(* Logix 5000 project; controller FV vendor 1 type 14 code 217 rev 31.11; software revision 31.00; part 41 of 63 *)
(* tags used below, declared in another part *)
   CWD : CHECKWORD_FLAGS;
   FV_AV1 : PlantItem;   // AV1
   FV_B100 : INT[255];   // FV FLAGS
   FV_B22 : INT[255];   // YSVFILL_FL YSV filling process flags
   FV_B22_0_2_OutputBit : BOOL;
   fv_data_file_value_to_move : DINT;
   FV_indirect_address : DINT;
   FV_N101 : INT[255];   // FV INT Fermentation control integer workspace
   FV_N104 : INT[255];   // FV_PC_BUF PC>PLC Fermentation Control Command Buff er File
   FV_N12 : INT[255];   // SYS_PARMS System Parameter Fil e
   FV_N141 : INT[255];   // YSV1 DATA
   FV_N142 : INT[255];   // YSV2 DATA
   FV_N143 : INT[255];   // YSV3 DATA
   FV_N144 : INT[255];   // YST1 DATA
   FV_N145 : INT[255];   // YST2 DATA
   FV_N20 : INT[255];   // YSVFILL<PC YSV Filling data fro m PC
   FV_N21 : INT[255];   // YSVFILL>PC YSV Filling process data to PC and contr ol regs
   FV_N24 : INT[255];   // YSVFILL_SV YSV filling process data save file to PC
   FV_YSV2O : PlantItem;   // YSV2O
   FV_YSV3O : PlantItem;   // YSV3O
   indirect_bit_temp : INT;
   YSVFilling_transaction_log_delay : DINT;
(* FV_Common, continued *)

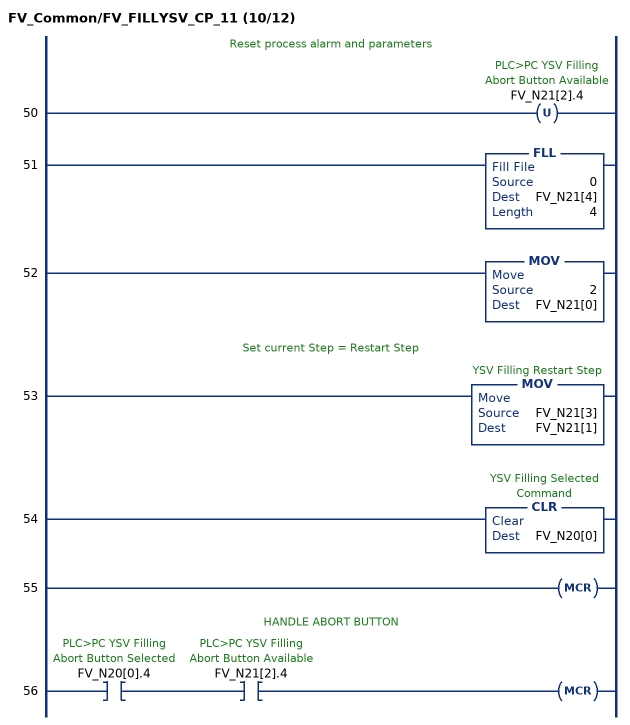
   // Reset process alarm and parameters
   50: OTU(FV_N21[2].4);
   51: FLL(0,FV_N21[4],4);
   52: MOV(2,FV_N21[0]);
   // Set current Step = Restart Step
   53: MOV(FV_N21[3],FV_N21[1]);
   54: CLR(FV_N20[0]);
   55: MCR();
   // HANDLE ABORT BUTTON
   56: XIC(FV_N20[0].4)XIC(FV_N21[2].4)MCR();
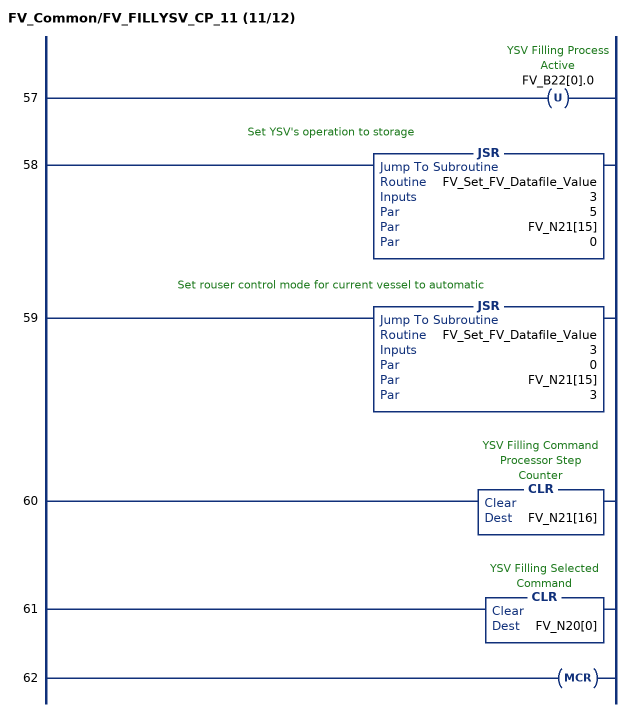
   57: OTU(FV_B22[0].0);
   // Set YSV's operation to storage
   58: JSR(FV_Set_FV_Datafile_Value,3,5,FV_N21[15],0);
   // Set rouser control mode for current vessel to automatic
   59: JSR(FV_Set_FV_Datafile_Value,3,0,FV_N21[15],3);
   60: CLR(FV_N21[16]);
   61: CLR(FV_N20[0]);
   62: MCR();
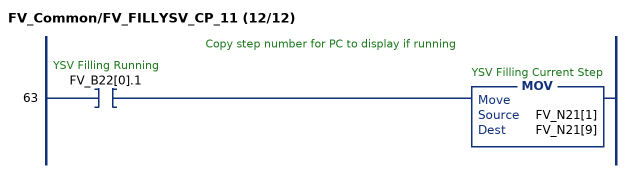
   // Copy step number for PC to display if running
   63: XIC(FV_B22[0].1)MOV(FV_N21[1],FV_N21[9]);
END_ROUTINE

ROUTINE FV_FILLYSV_MC_10   (* ladder *)
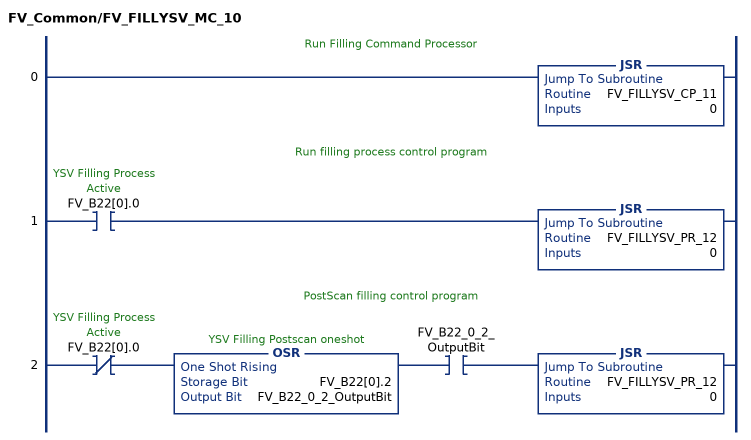
   // Run Filling Command Processor
   0: JSR(FV_FILLYSV_CP_11,0);
   // Run filling process control program
   1: XIC(FV_B22[0].0)JSR(FV_FILLYSV_PR_12,0);
   // PostScan filling control program
   2: XIO(FV_B22[0].0)OSR(FV_B22[0].2,FV_B22_0_2_OutputBit)XIC(FV_B22_0_2_OutputBit)JSR(FV_FILLYSV_PR_12,0);
END_ROUTINE

ROUTINE FV_FILLYSV_PR_12   (* ladder *)
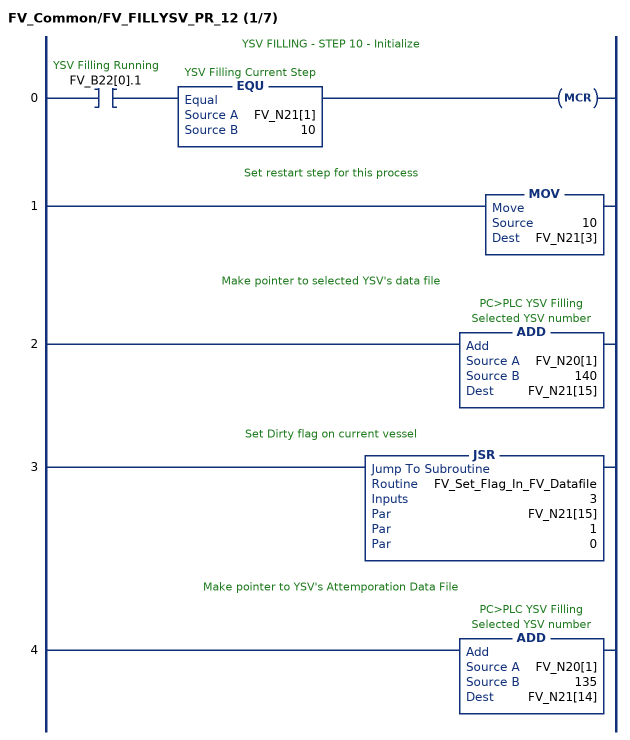
   // YSV FILLING - STEP 10 - Initialize
   0: XIC(FV_B22[0].1)EQU(FV_N21[1],10)MCR();
   // Set restart step for this process
   1: MOV(10,FV_N21[3]);
   // Make pointer to selected YSV's data file
   2: ADD(FV_N20[1],140,FV_N21[15]);
   // Set Dirty flag on current vessel
   3: JSR(FV_Set_Flag_In_FV_Datafile,3,FV_N21[15],1,0);
   // Make pointer to YSV's Attemporation Data File
   4: ADD(FV_N20[1],135,FV_N21[14]);
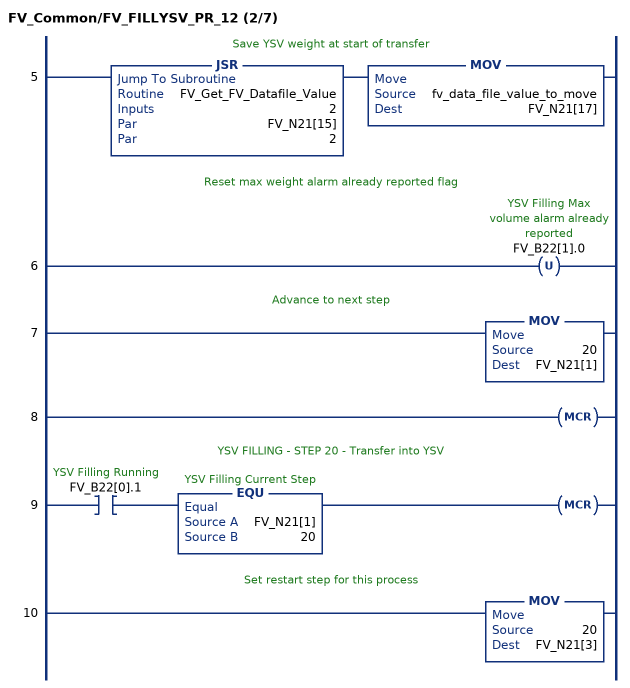
   // Save YSV weight at start of transfer
   5: JSR(FV_Get_FV_Datafile_Value,2,FV_N21[15],2)MOV(fv_data_file_value_to_move,FV_N21[17]);
   // Reset max weight alarm already reported flag
   6: OTU(FV_B22[1].0);
   // Advance to next step
   7: MOV(20,FV_N21[1]);
   8: MCR();
   // YSV FILLING - STEP 20 - Transfer into YSV
   9: XIC(FV_B22[0].1)EQU(FV_N21[1],20)MCR();
   // Set restart step for this process
   10: MOV(20,FV_N21[3]);
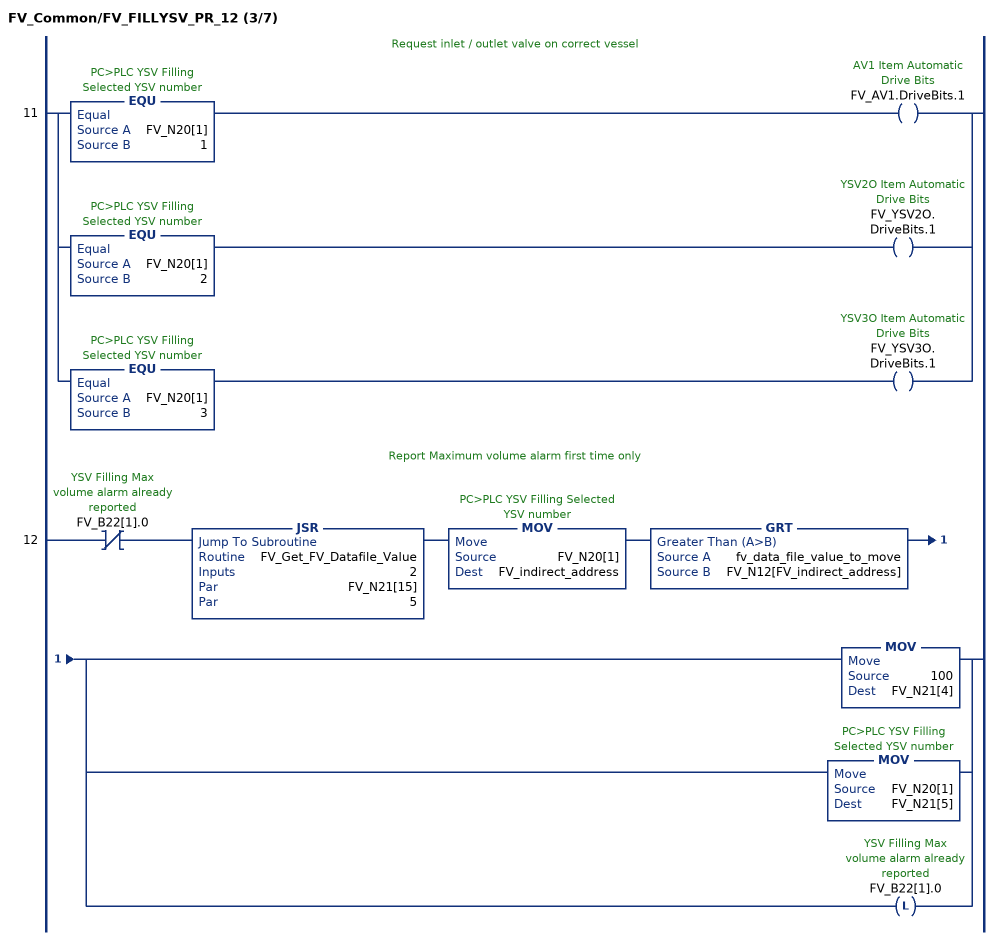
   // Request inlet / outlet valve on correct vessel
   11: [EQU(FV_N20[1],1) OTE(FV_AV1.DriveBits.1) ,EQU(FV_N20[1],2) OTE(FV_YSV2O.DriveBits.1) ,EQU(FV_N20[1],3) OTE(FV_YSV3O.DriveBits.1) ];
   // Report Maximum volume alarm first time only
   12: XIO(FV_B22[1].0)JSR(FV_Get_FV_Datafile_Value,2,FV_N21[15],5)MOV(FV_N20[1],FV_indirect_address)GRT(fv_data_file_value_to_move,FV_N12[FV_indirect_address])[MOV(100,FV_N21[4]) ,MOV(FV_N20[1],FV_N21[5]) ,OTL(FV_B22[1].0) ];
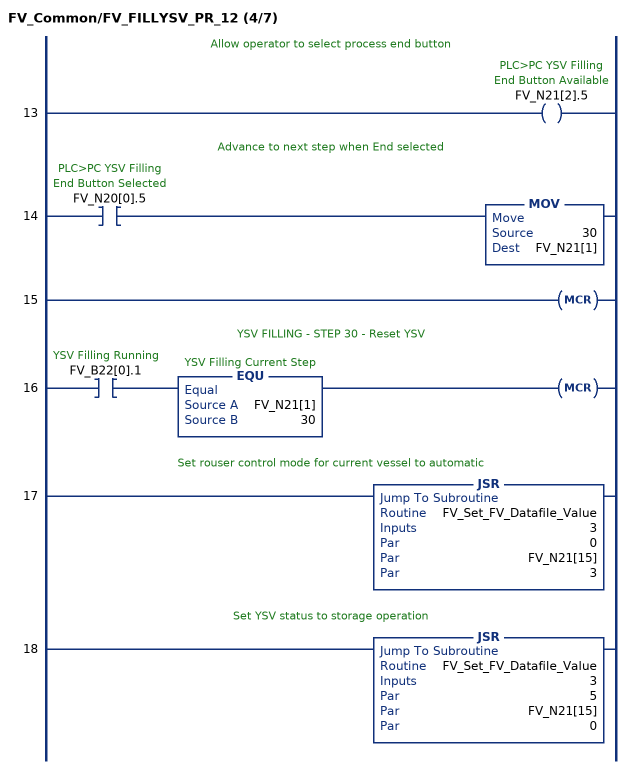
   // Allow operator to select process end button
   13: OTE(FV_N21[2].5);
   // Advance to next step when End selected
   14: XIC(FV_N20[0].5)MOV(30,FV_N21[1]);
   15: MCR();
   // YSV FILLING - STEP 30 - Reset YSV
   16: XIC(FV_B22[0].1)EQU(FV_N21[1],30)MCR();
   // Set rouser control mode for current vessel to automatic
   17: JSR(FV_Set_FV_Datafile_Value,3,0,FV_N21[15],3);
   // Set YSV status to storage operation
   18: JSR(FV_Set_FV_Datafile_Value,3,5,FV_N21[15],0);
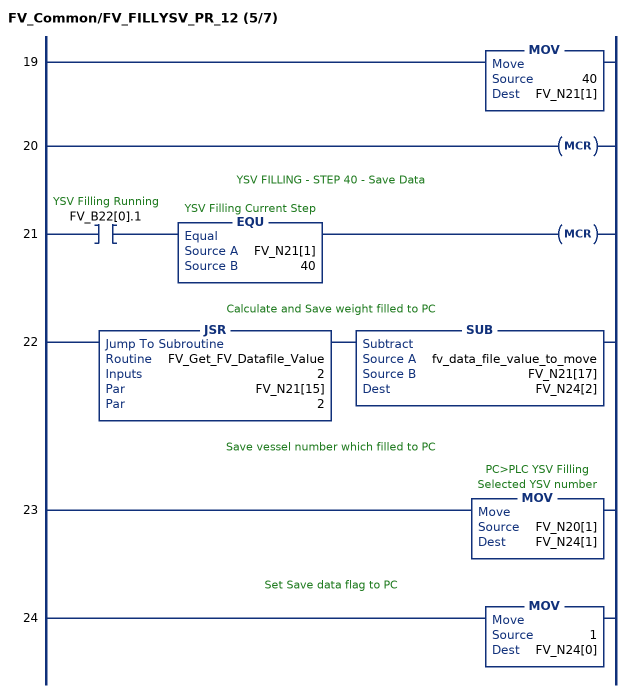
   19: MOV(40,FV_N21[1]);
   20: MCR();
   // YSV FILLING - STEP 40 - Save Data
   21: XIC(FV_B22[0].1)EQU(FV_N21[1],40)MCR();
   // Calculate and Save weight filled to PC
   22: JSR(FV_Get_FV_Datafile_Value,2,FV_N21[15],2)SUB(fv_data_file_value_to_move,FV_N21[17],FV_N24[2]);
   // Save vessel number which filled to PC
   23: MOV(FV_N20[1],FV_N24[1]);
   // Set Save data flag to PC
   24: MOV(1,FV_N24[0]);
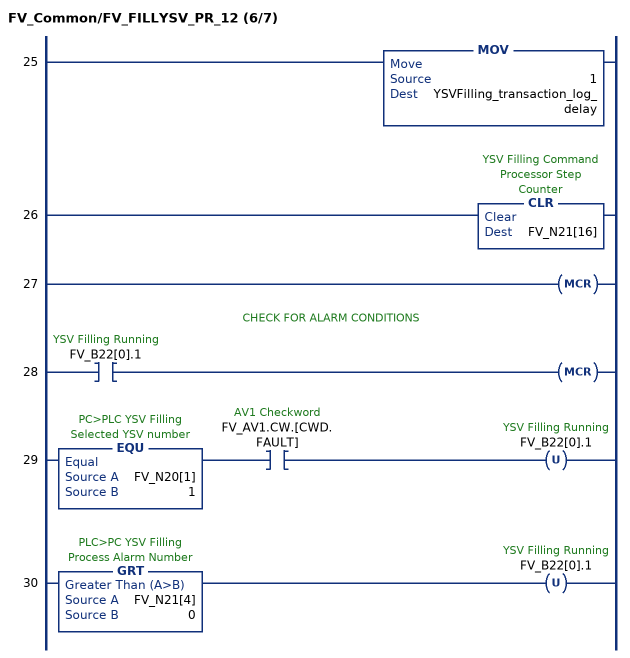
   25: MOV(1,YSVFilling_transaction_log_delay);
   26: CLR(FV_N21[16]);
   27: MCR();
   // CHECK FOR ALARM CONDITIONS
   28: XIC(FV_B22[0].1)MCR();
   29: EQU(FV_N20[1],1)XIC(FV_AV1.CW.[CWD.FAULT])OTU(FV_B22[0].1);
   30: GRT(FV_N21[4],0)OTU(FV_B22[0].1);
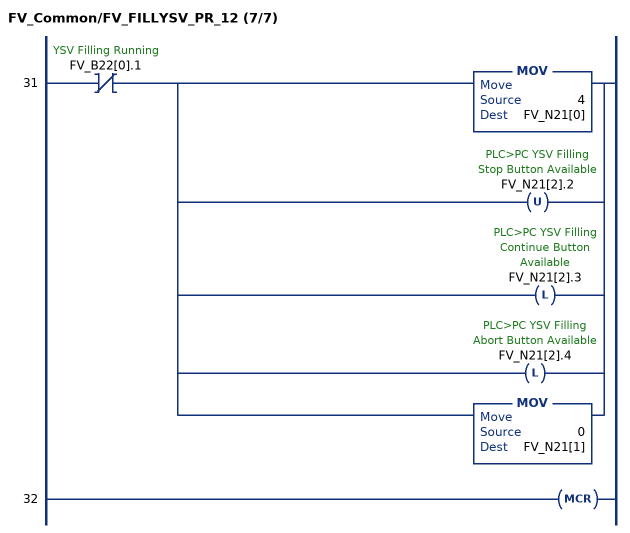
   31: XIO(FV_B22[0].1)[MOV(4,FV_N21[0]) ,OTU(FV_N21[2].2) ,OTL(FV_N21[2].3) ,OTL(FV_N21[2].4) ,MOV(0,FV_N21[1]) ];
   32: MCR();
END_ROUTINE

ROUTINE FV_FV_COMMAND_101   (* ladder *)
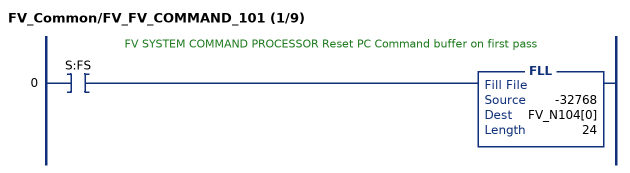
   // FV SYSTEM COMMAND PROCESSOR Reset PC Command buffer on first pass
   0: XIC(S:FS)FLL(-32768,FV_N104[0],24);
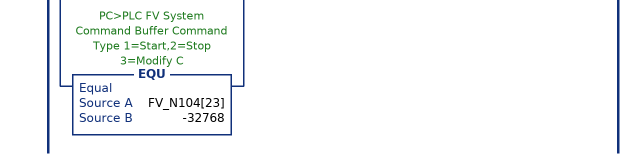
   // WAIT FOR PC TO SEND NEW FV SYSTEM COMMAND If any word within the PC/PLC FV system command buffer contains -32768, the block has not yet been fully downloaded and therefore no new command has been requested.
   1: [EQU(FV_N104[0],-32768) ,EQU(FV_N104[1],-32768) ,EQU(FV_N104[2],-32768) ,EQU(FV_N104[3],-32768) ,EQU(FV_N104[4],-32768) ,EQU(FV_N104[5],-32768) ,EQU(FV_N104[6],-32768) ,EQU(FV_N104[7],-32768) ,EQU(FV_N104[8],-32768) ,EQU(FV_N104[9],-32768) ,EQU(FV_N104[10],-32768) ,EQU(FV_N104[11],-32768) ,EQU(FV_N104[12],-32768) ,EQU(FV_N104[13],-32768) ,EQU(FV_N104[14],-32768) ,EQU(FV_N104[15],-32768) ,EQU(FV_N104[16],-32768) ,EQU(FV_N104[17],-32768) ,EQU(FV_N104[18],-32768) ,EQU(FV_N104[19],-32768) ,EQU(FV_N104[20],-32768) ,EQU(FV_N104[21],-32768) ,EQU(FV_N104[22],-32768) ,EQU(FV_N104[23],-32768) ]OTE(FV_B100[1].0);
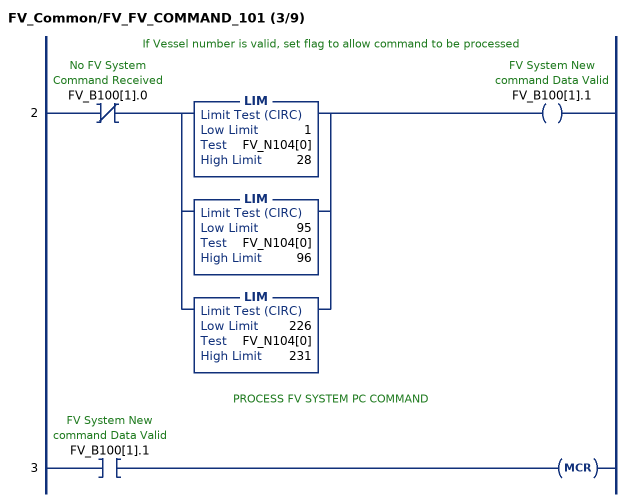
   // If Vessel number is valid, set flag to allow command to be processed
   2: XIO(FV_B100[1].0)[LIM(1,FV_N104[0],28) ,LIM(95,FV_N104[0],96) ,LIM(226,FV_N104[0],231) ]OTE(FV_B100[1].1);
   // PROCESS FV SYSTEM PC COMMAND
   3: XIC(FV_B100[1].1)MCR();
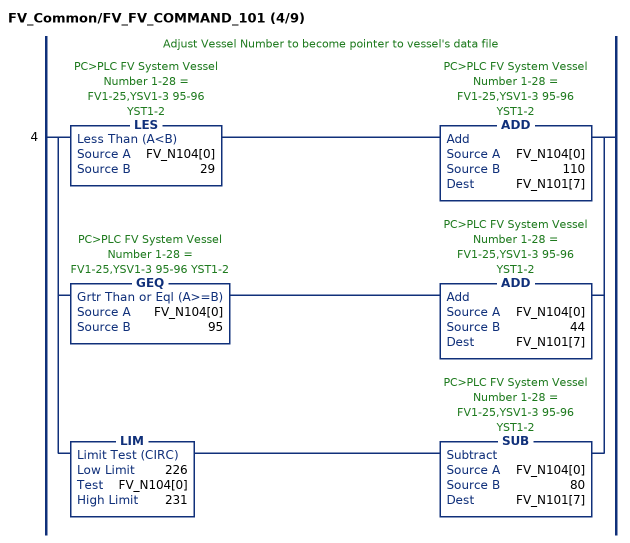
   // Adjust Vessel Number to become pointer to vessel's data file
   4: [LES(FV_N104[0],29) ADD(FV_N104[0],110,FV_N101[7]) ,GEQ(FV_N104[0],95) ADD(FV_N104[0],44,FV_N101[7]) ,LIM(226,FV_N104[0],231) SUB(FV_N104[0],80,FV_N101[7]) ];
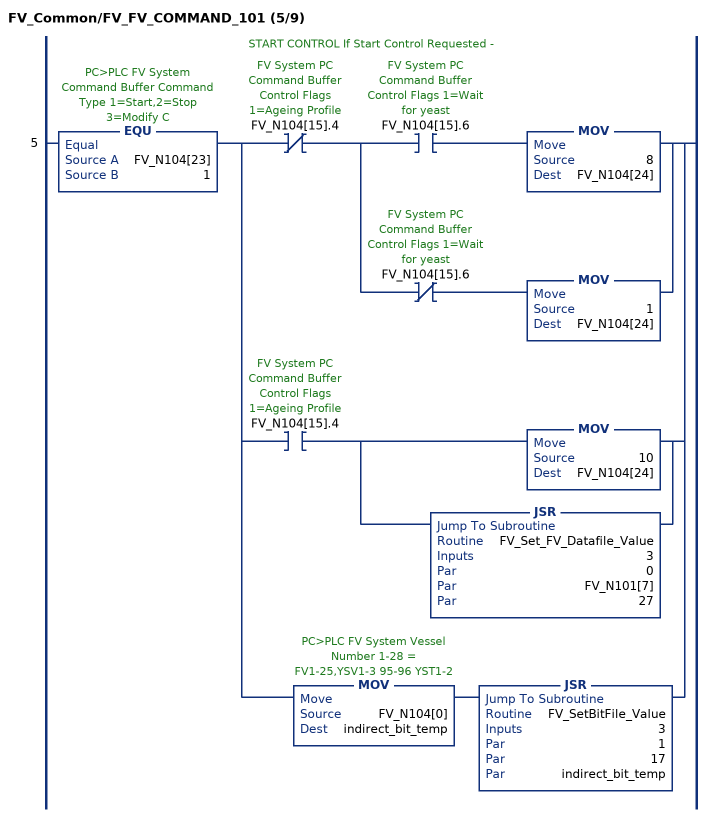
   // START CONTROL If Start Control Requested -
   5: EQU(FV_N104[23],1)[XIO(FV_N104[15].4) [XIC(FV_N104[15].6) MOV(8,FV_N104[24]) ,XIO(FV_N104[15].6) MOV(1,FV_N104[24]) ] ,XIC(FV_N104[15].4) [MOV(10,FV_N104[24]) ,JSR(FV_Set_FV_Datafile_Value,3,0,FV_N101[7],27) ] ,MOV(FV_N104[0],indirect_bit_temp) JSR(FV_SetBitFile_Value,3,1,17,indirect_bit_temp) ];
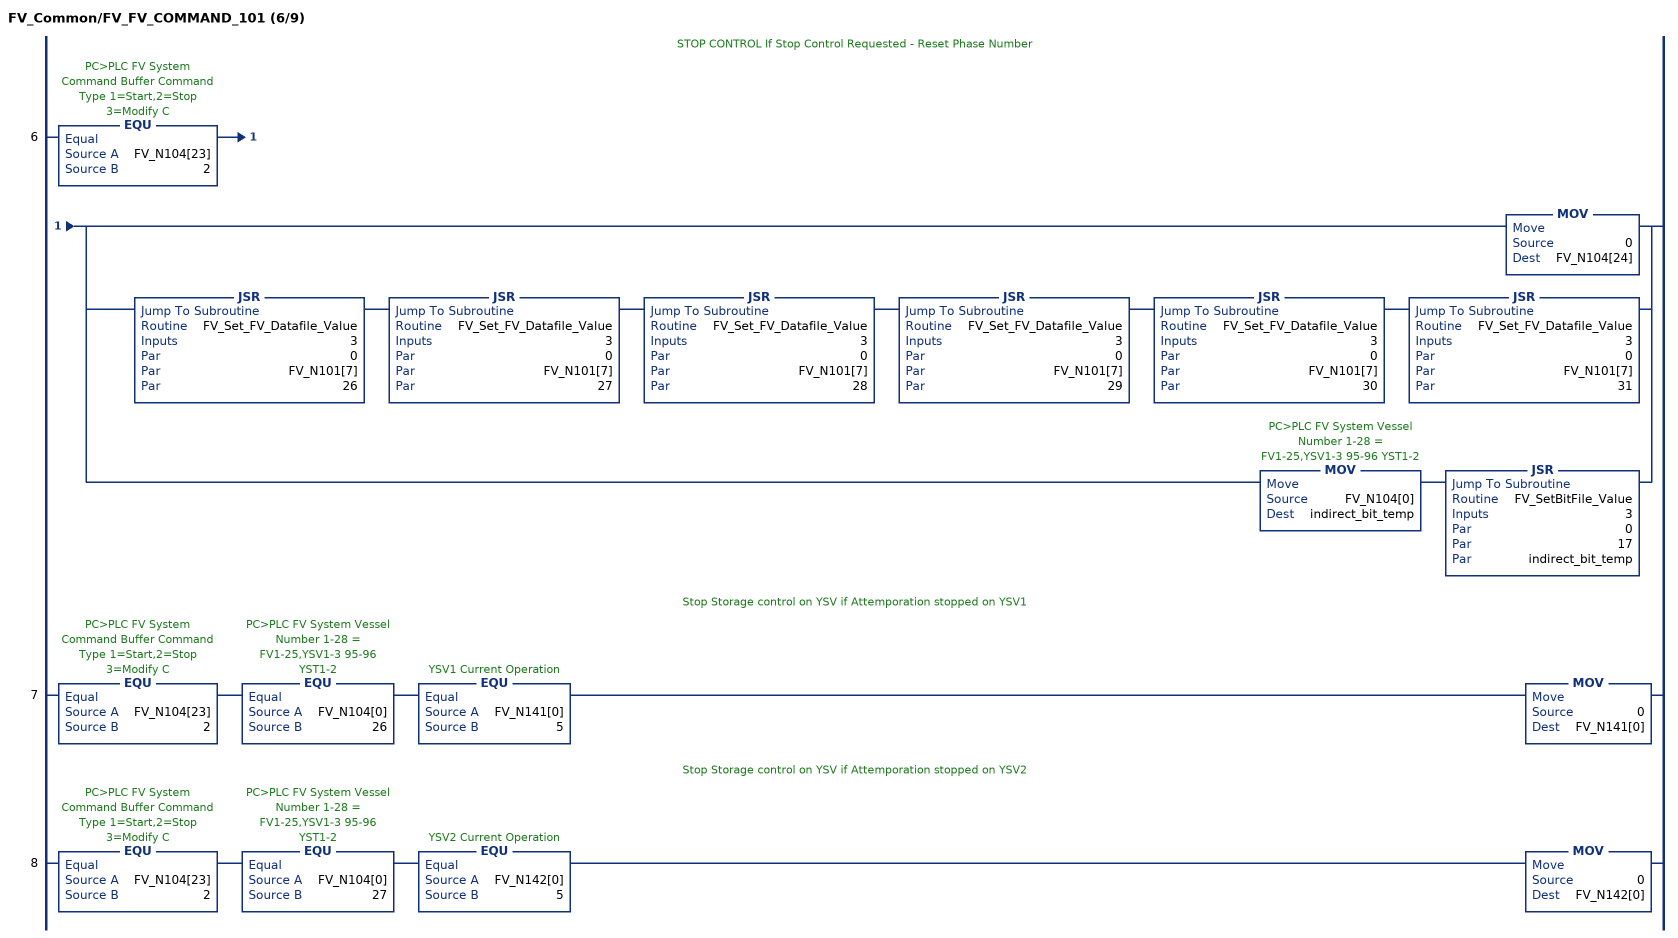
   // STOP CONTROL If Stop Control Requested - Reset Phase Number
   6: EQU(FV_N104[23],2)[MOV(0,FV_N104[24]) ,JSR(FV_Set_FV_Datafile_Value,3,0,FV_N101[7],26) JSR(FV_Set_FV_Datafile_Value,3,0,FV_N101[7],27) JSR(FV_Set_FV_Datafile_Value,3,0,FV_N101[7],28) JSR(FV_Set_FV_Datafile_Value,3,0,FV_N101[7],29) JSR(FV_Set_FV_Datafile_Value,3,0,FV_N101[7],30) JSR(FV_Set_FV_Datafile_Value,3,0,FV_N101[7],31) ,MOV(FV_N104[0],indirect_bit_temp) JSR(FV_SetBitFile_Value,3,0,17,indirect_bit_temp) ];
   // Stop Storage control on YSV if Attemporation stopped on YSV1
   7: EQU(FV_N104[23],2)EQU(FV_N104[0],26)EQU(FV_N141[0],5)MOV(0,FV_N141[0]);
   // Stop Storage control on YSV if Attemporation stopped on YSV2
   8: EQU(FV_N104[23],2)EQU(FV_N104[0],27)EQU(FV_N142[0],5)MOV(0,FV_N142[0]);
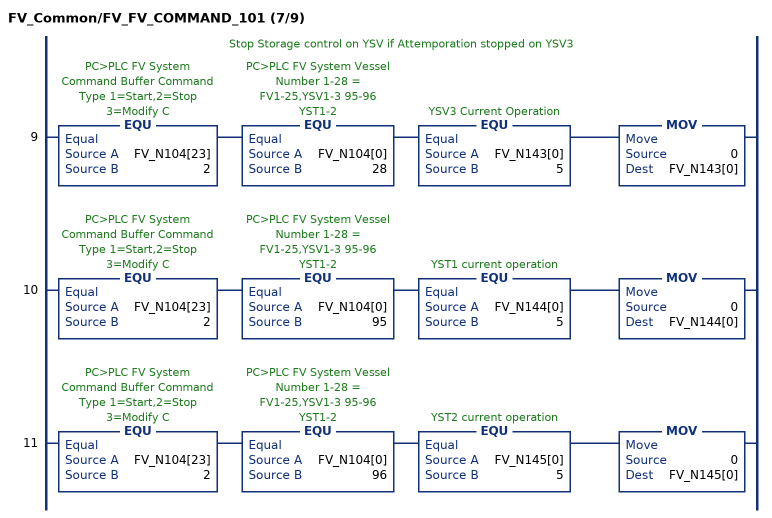
   // Stop Storage control on YSV if Attemporation stopped on YSV3
   9: EQU(FV_N104[23],2)EQU(FV_N104[0],28)EQU(FV_N143[0],5)MOV(0,FV_N143[0]);
   10: EQU(FV_N104[23],2)EQU(FV_N104[0],95)EQU(FV_N144[0],5)MOV(0,FV_N144[0]);
   11: EQU(FV_N104[23],2)EQU(FV_N104[0],96)EQU(FV_N145[0],5)MOV(0,FV_N145[0]);
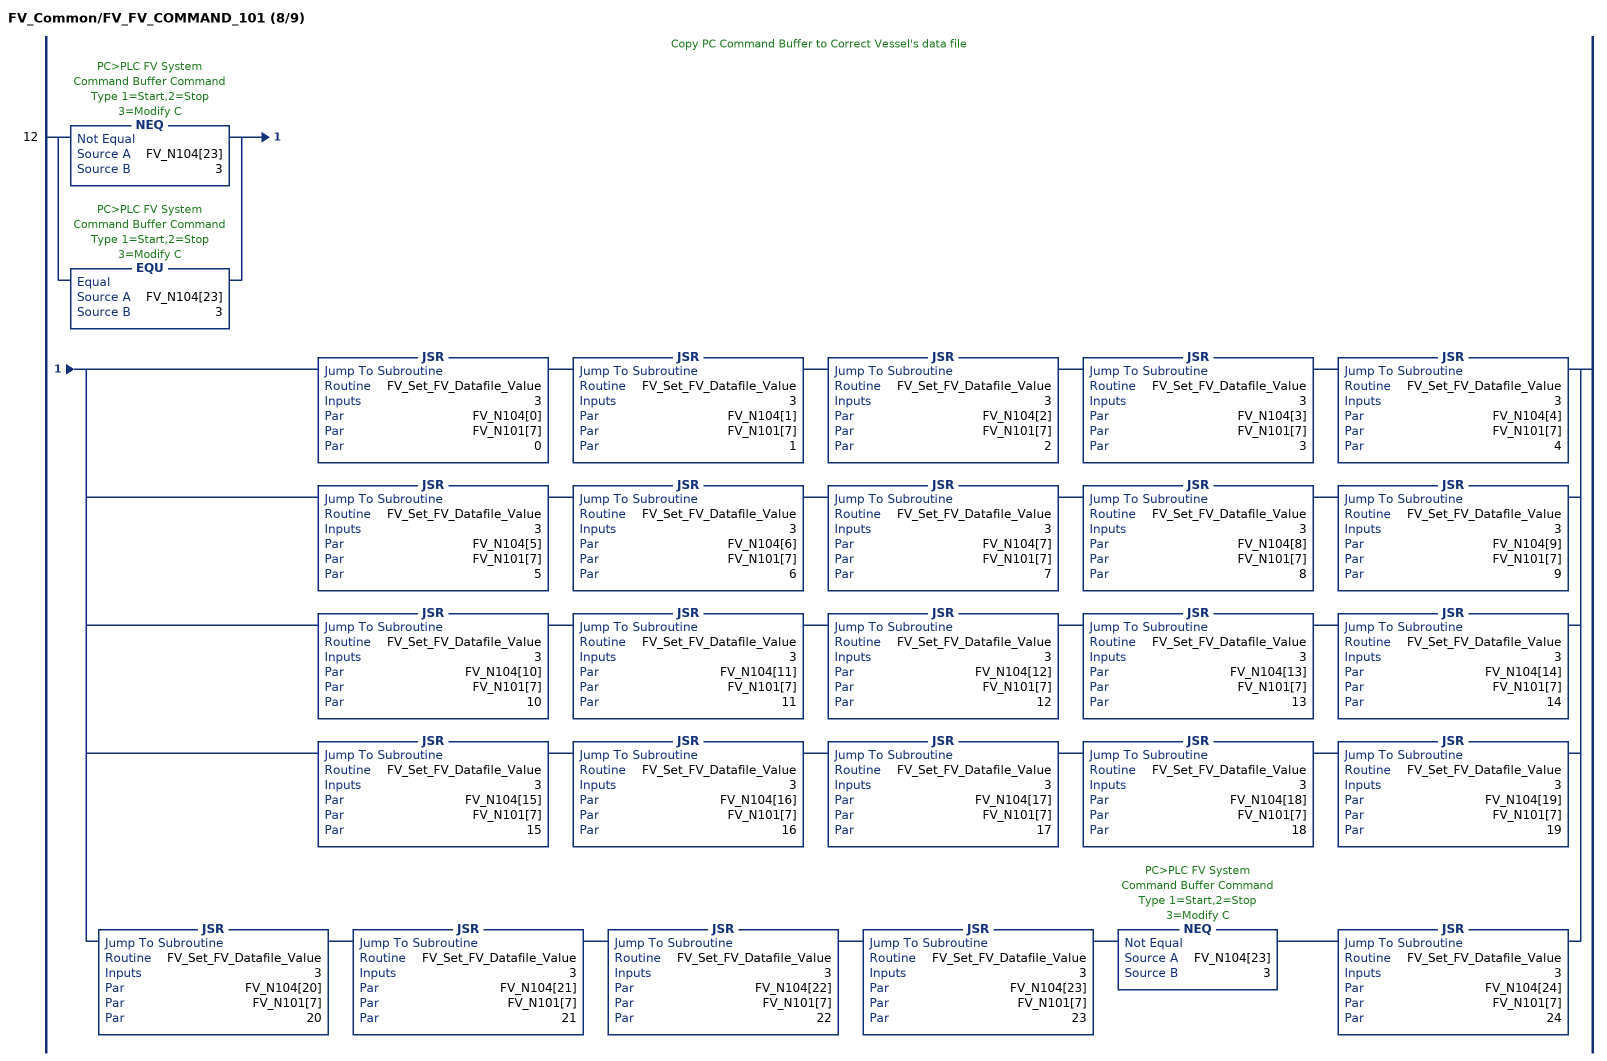
   // Copy PC Command Buffer to Correct Vessel's data file
   12: [NEQ(FV_N104[23],3) ,EQU(FV_N104[23],3) ][JSR(FV_Set_FV_Datafile_Value,3,FV_N104[0],FV_N101[7],0) JSR(FV_Set_FV_Datafile_Value,3,FV_N104[1],FV_N101[7],1) JSR(FV_Set_FV_Datafile_Value,3,FV_N104[2],FV_N101[7],2) JSR(FV_Set_FV_Datafile_Value,3,FV_N104[3],FV_N101[7],3) JSR(FV_Set_FV_Datafile_Value,3,FV_N104[4],FV_N101[7],4) ,JSR(FV_Set_FV_Datafile_Value,3,FV_N104[5],FV_N101[7],5) JSR(FV_Set_FV_Datafile_Value,3,FV_N104[6],FV_N101[7],6) JSR(FV_Set_FV_Datafile_Value,3,FV_N104[7],FV_N101[7],7) JSR(FV_Set_FV_Datafile_Value,3,FV_N104[8],FV_N101[7],8) JSR(FV_Set_FV_Datafile_Value,3,FV_N104[9],FV_N101[7],9) ,JSR(FV_Set_FV_Datafile_Value,3,FV_N104[10],FV_N101[7],10) JSR(FV_Set_FV_Datafile_Value,3,FV_N104[11],FV_N101[7],11) JSR(FV_Set_FV_Datafile_Value,3,FV_N104[12],FV_N101[7],12) JSR(FV_Set_FV_Datafile_Value,3,FV_N104[13],FV_N101[7],13) JSR(FV_Set_FV_Datafile_Value,3,FV_N104[14],FV_N101[7],14) ,JSR(FV_Set_FV_Datafile_Value,3,FV_N104[15],FV_N101[7],15) JSR(FV_Set_FV_Datafile_Value,3,FV_N104[16],FV_N101[7],16) JSR(FV_Set_FV_Datafile_Value,3,FV_N104[17],FV_N101[7],17) JSR(FV_Set_FV_Datafile_Value,3,FV_N104[18],FV_N101[7],18) JSR(FV_Set_FV_Datafile_Value,3,FV_N104[19],FV_N101[7],19) ,JSR(FV_Set_FV_Datafile_Value,3,FV_N104[20],FV_N101[7],20) JSR(FV_Set_FV_Datafile_Value,3,FV_N104[21],FV_N101[7],21) JSR(FV_Set_FV_Datafile_Value,3,FV_N104[22],FV_N101[7],22) JSR(FV_Set_FV_Datafile_Value,3,FV_N104[23],FV_N101[7],23) NEQ(FV_N104[23],3) JSR(FV_Set_FV_Datafile_Value,3,FV_N104[24],FV_N101[7],24) ];
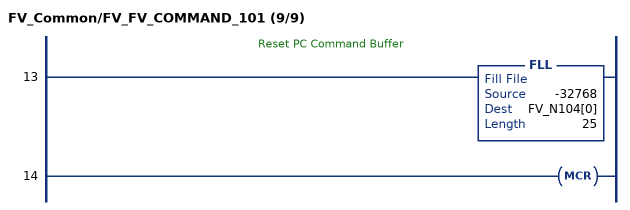
   // Reset PC Command Buffer
   13: FLL(-32768,FV_N104[0],25);
   14: MCR();
END_ROUTINE
